(* Logix 5000 project; controller FV vendor 1 type 14 code 217 rev 31.11; software revision 31.00; part 10 of 63 *)
(* tags used below, declared in another part *)
   CWD : CHECKWORD_FLAGS;
   FR_AUDI1 : PlantItem;   // AUDI1
   FR_AUDI1_RawOutput : ALIAS FOR RIO_Rack_2:11:O.Data.30;   // FR_AUDI1
   FR_BEACON1 : PlantItem;   // BEACON1
   FR_BEACON1_RawOutput : ALIAS FOR RIO_Rack_2:11:O.Data.31;   // FR_BEACON1
   FR_data_file_value_to_move : DINT;
   FR_DEFOAM : PlantItem;   // DEFOAM
   FR_DEFOAM_RawOutput : ALIAS FOR RIO_Rack_2:5:O.Data.6;   // FR_DEFOAM
   FR_Delphi_O : DINT[60];
   FR_FV26_VA01 : PlantItem;   // FV26_VA01
   FR_FV26_VA01_RawOutput : ALIAS FOR RIO_Rack_2:11:O.Data.24;   // FR_FV26_VA01
   FR_FV27_VA01 : PlantItem;   // FV27_VA01
   FR_FV27_VA01_RawOutput : ALIAS FOR RIO_Rack_2:11:O.Data.25;   // FR_FV27_VA01
   FR_FV28_V : PlantItem;   // FV28_V
   FR_FV28_V_RawOutput : ALIAS FOR RIO_Rack_2:11:O.Data.20;   // FR_FV28_V
   FR_FV28_VA01 : PlantItem;   // FV28_VA01
   FR_FV28_VA01_RawOutput : ALIAS FOR RIO_Rack_2:11:O.Data.26;   // FR_FV28_VA01
   FR_FV29_VA01 : PlantItem;   // FV29_VA01
   FR_FV29_VA01_RawOutput : ALIAS FOR RIO_Rack_2:11:O.Data.27;   // FR_FV29_VA01
   FR_FV30_VA01 : PlantItem;   // FV30_VA01
   FR_FV30_VA01_RawOutput : ALIAS FOR RIO_Rack_2:11:O.Data.28;   // FR_FV30_VA01
   FR_FV31_VA01 : PlantItem;   // FV31_VA01
   FR_FV31_VA01_RawOutput : ALIAS FOR RIO_Rack_2:11:O.Data.29;   // FR_FV31_VA01
   FR_FVR1_P01 : PlantItem;   // FVR1_P01
   FR_N130 : INT[265];   // FILTRATE Filtrate Return
   FR_N14 : INT[265];   // MVFV CIP Comms to MVFV CIP Un it PLC
   FR_N140 : INT[265];   // CIP
   FR_N160 : INT[265];   // VESSEL Vessel Working Direc tory
   FR_N99 : INT[265];   // COMMENT Comment Lines
   FR_T131 : TIMER[255];   // FILTRATE
   FR_T4 : TIMER[255];   // TIMER
   FR_YC_1 : PlantItem;   // YC_1
   FR_YC_1_RawOutput : ALIAS FOR RIO_Rack_2:11:O.Data.16;   // FR_YC_1
   FR_YC_2 : PlantItem;   // YC_2
   FR_YC_2_RawOutput : ALIAS FOR RIO_Rack_2:11:O.Data.17;   // FR_YC_2
   FR_YP1_CIP : PlantItem;   // YP1_CIP
   FR_YP1_CIP_RawOutput : ALIAS FOR RIO_Rack_2:11:O.Data.21;   // FR_YP1_CIP
   FR_YP2_CIP : PlantItem;   // YP2_CIP
   FR_YP2_CIP_RawOutput : ALIAS FOR RIO_Rack_2:11:O.Data.22;   // FR_YP2_CIP
   FR_YP3_CIP : PlantItem;   // YP3_CIP
   FR_YP3_CIP_RawOutput : ALIAS FOR RIO_Rack_2:11:O.Data.23;   // FR_YP3_CIP
   FT_Filtrate_131_temp_real : REAL;
(* FR_Common, continued *)

ROUTINE FR_Digital_Outputs   (* ladder *)
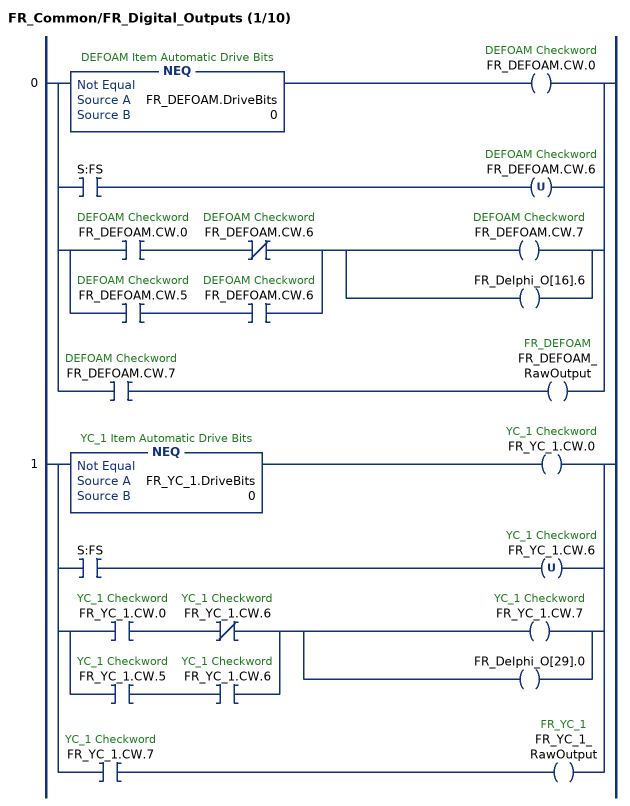
   0: [NEQ(FR_DEFOAM.DriveBits,0) OTE(FR_DEFOAM.CW.0) ,XIC(S:FS) OTU(FR_DEFOAM.CW.6) ,[XIC(FR_DEFOAM.CW.0) XIO(FR_DEFOAM.CW.6) ,XIC(FR_DEFOAM.CW.5) XIC(FR_DEFOAM.CW.6) ] [OTE(FR_DEFOAM.CW.7) ,OTE(FR_Delphi_O[16].6) ] ,XIC(FR_DEFOAM.CW.7) OTE(FR_DEFOAM_RawOutput) ];
   1: [NEQ(FR_YC_1.DriveBits,0) OTE(FR_YC_1.CW.0) ,XIC(S:FS) OTU(FR_YC_1.CW.6) ,[XIC(FR_YC_1.CW.0) XIO(FR_YC_1.CW.6) ,XIC(FR_YC_1.CW.5) XIC(FR_YC_1.CW.6) ] [OTE(FR_YC_1.CW.7) ,OTE(FR_Delphi_O[29].0) ] ,XIC(FR_YC_1.CW.7) OTE(FR_YC_1_RawOutput) ];
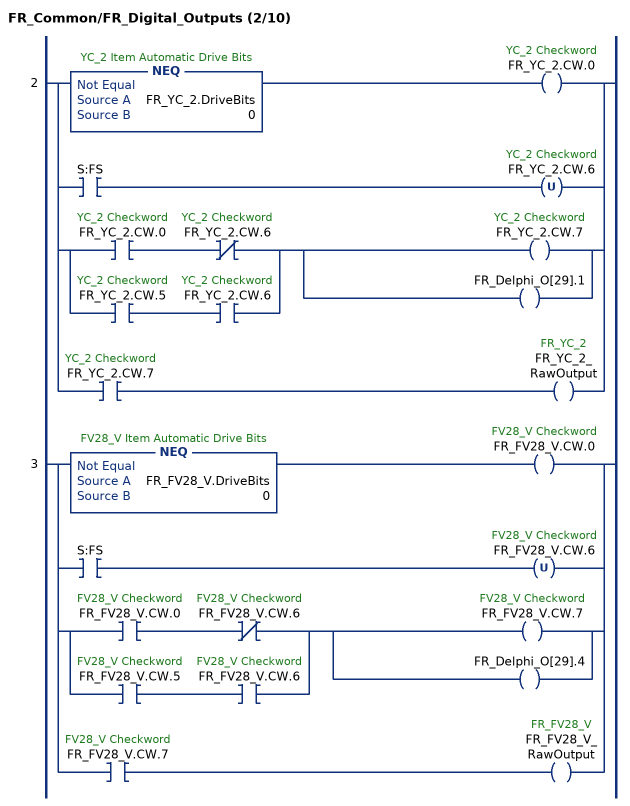
   2: [NEQ(FR_YC_2.DriveBits,0) OTE(FR_YC_2.CW.0) ,XIC(S:FS) OTU(FR_YC_2.CW.6) ,[XIC(FR_YC_2.CW.0) XIO(FR_YC_2.CW.6) ,XIC(FR_YC_2.CW.5) XIC(FR_YC_2.CW.6) ] [OTE(FR_YC_2.CW.7) ,OTE(FR_Delphi_O[29].1) ] ,XIC(FR_YC_2.CW.7) OTE(FR_YC_2_RawOutput) ];
   3: [NEQ(FR_FV28_V.DriveBits,0) OTE(FR_FV28_V.CW.0) ,XIC(S:FS) OTU(FR_FV28_V.CW.6) ,[XIC(FR_FV28_V.CW.0) XIO(FR_FV28_V.CW.6) ,XIC(FR_FV28_V.CW.5) XIC(FR_FV28_V.CW.6) ] [OTE(FR_FV28_V.CW.7) ,OTE(FR_Delphi_O[29].4) ] ,XIC(FR_FV28_V.CW.7) OTE(FR_FV28_V_RawOutput) ];
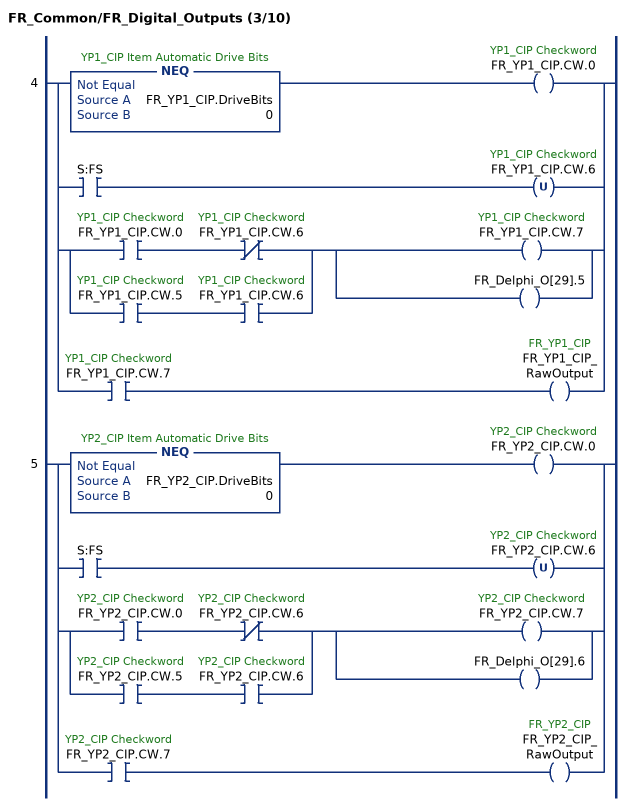
   4: [NEQ(FR_YP1_CIP.DriveBits,0) OTE(FR_YP1_CIP.CW.0) ,XIC(S:FS) OTU(FR_YP1_CIP.CW.6) ,[XIC(FR_YP1_CIP.CW.0) XIO(FR_YP1_CIP.CW.6) ,XIC(FR_YP1_CIP.CW.5) XIC(FR_YP1_CIP.CW.6) ] [OTE(FR_YP1_CIP.CW.7) ,OTE(FR_Delphi_O[29].5) ] ,XIC(FR_YP1_CIP.CW.7) OTE(FR_YP1_CIP_RawOutput) ];
   5: [NEQ(FR_YP2_CIP.DriveBits,0) OTE(FR_YP2_CIP.CW.0) ,XIC(S:FS) OTU(FR_YP2_CIP.CW.6) ,[XIC(FR_YP2_CIP.CW.0) XIO(FR_YP2_CIP.CW.6) ,XIC(FR_YP2_CIP.CW.5) XIC(FR_YP2_CIP.CW.6) ] [OTE(FR_YP2_CIP.CW.7) ,OTE(FR_Delphi_O[29].6) ] ,XIC(FR_YP2_CIP.CW.7) OTE(FR_YP2_CIP_RawOutput) ];
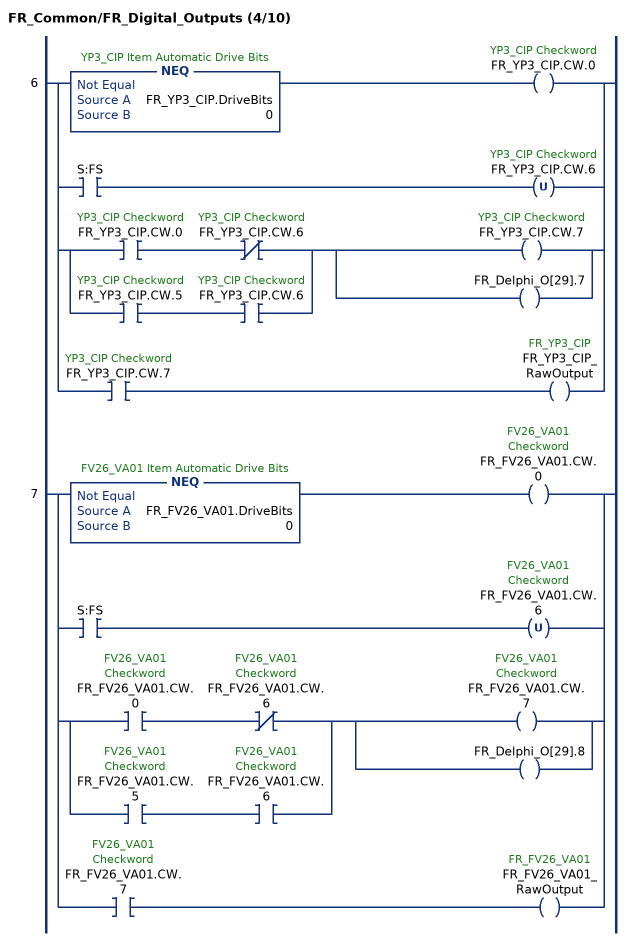
   6: [NEQ(FR_YP3_CIP.DriveBits,0) OTE(FR_YP3_CIP.CW.0) ,XIC(S:FS) OTU(FR_YP3_CIP.CW.6) ,[XIC(FR_YP3_CIP.CW.0) XIO(FR_YP3_CIP.CW.6) ,XIC(FR_YP3_CIP.CW.5) XIC(FR_YP3_CIP.CW.6) ] [OTE(FR_YP3_CIP.CW.7) ,OTE(FR_Delphi_O[29].7) ] ,XIC(FR_YP3_CIP.CW.7) OTE(FR_YP3_CIP_RawOutput) ];
   7: [NEQ(FR_FV26_VA01.DriveBits,0) OTE(FR_FV26_VA01.CW.0) ,XIC(S:FS) OTU(FR_FV26_VA01.CW.6) ,[XIC(FR_FV26_VA01.CW.0) XIO(FR_FV26_VA01.CW.6) ,XIC(FR_FV26_VA01.CW.5) XIC(FR_FV26_VA01.CW.6) ] [OTE(FR_FV26_VA01.CW.7) ,OTE(FR_Delphi_O[29].8) ] ,XIC(FR_FV26_VA01.CW.7) OTE(FR_FV26_VA01_RawOutput) ];
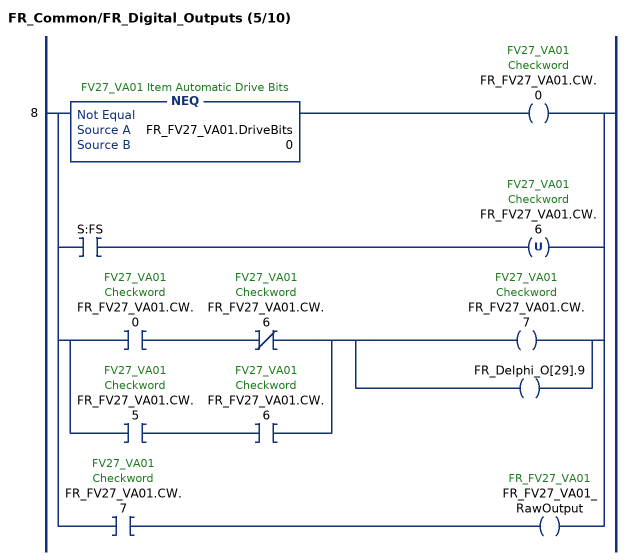
   8: [NEQ(FR_FV27_VA01.DriveBits,0) OTE(FR_FV27_VA01.CW.0) ,XIC(S:FS) OTU(FR_FV27_VA01.CW.6) ,[XIC(FR_FV27_VA01.CW.0) XIO(FR_FV27_VA01.CW.6) ,XIC(FR_FV27_VA01.CW.5) XIC(FR_FV27_VA01.CW.6) ] [OTE(FR_FV27_VA01.CW.7) ,OTE(FR_Delphi_O[29].9) ] ,XIC(FR_FV27_VA01.CW.7) OTE(FR_FV27_VA01_RawOutput) ];
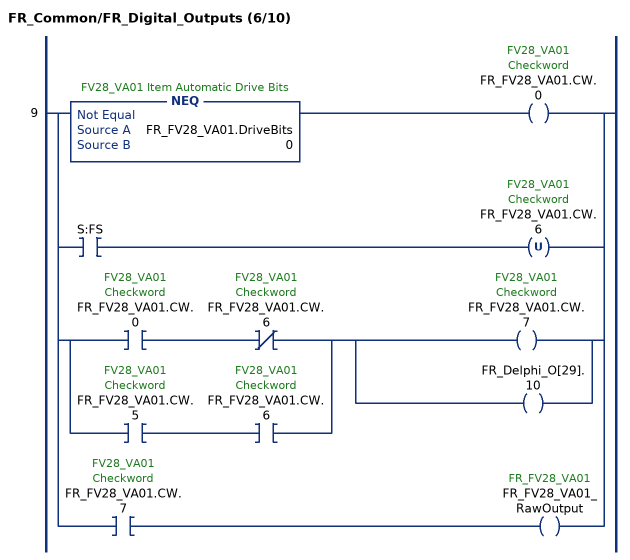
   9: [NEQ(FR_FV28_VA01.DriveBits,0) OTE(FR_FV28_VA01.CW.0) ,XIC(S:FS) OTU(FR_FV28_VA01.CW.6) ,[XIC(FR_FV28_VA01.CW.0) XIO(FR_FV28_VA01.CW.6) ,XIC(FR_FV28_VA01.CW.5) XIC(FR_FV28_VA01.CW.6) ] [OTE(FR_FV28_VA01.CW.7) ,OTE(FR_Delphi_O[29].10) ] ,XIC(FR_FV28_VA01.CW.7) OTE(FR_FV28_VA01_RawOutput) ];
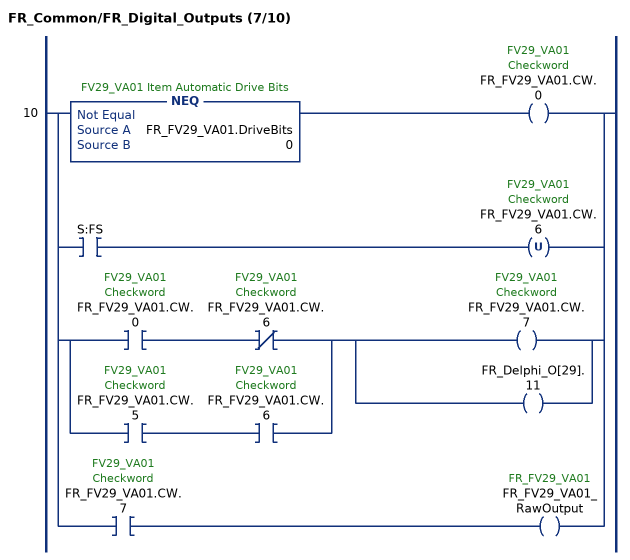
   10: [NEQ(FR_FV29_VA01.DriveBits,0) OTE(FR_FV29_VA01.CW.0) ,XIC(S:FS) OTU(FR_FV29_VA01.CW.6) ,[XIC(FR_FV29_VA01.CW.0) XIO(FR_FV29_VA01.CW.6) ,XIC(FR_FV29_VA01.CW.5) XIC(FR_FV29_VA01.CW.6) ] [OTE(FR_FV29_VA01.CW.7) ,OTE(FR_Delphi_O[29].11) ] ,XIC(FR_FV29_VA01.CW.7) OTE(FR_FV29_VA01_RawOutput) ];
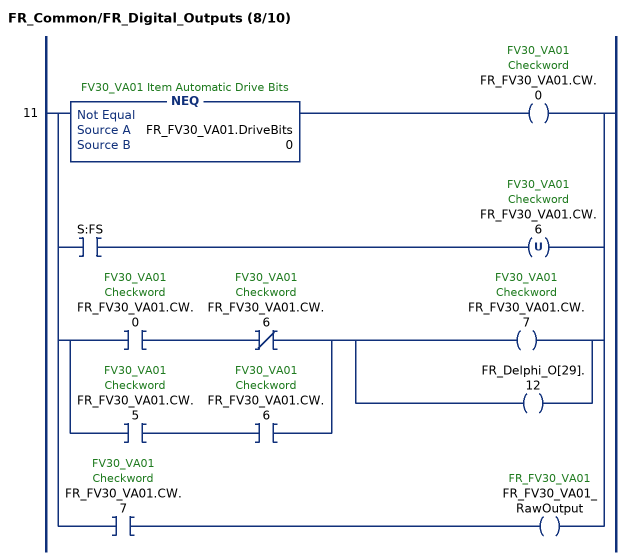
   11: [NEQ(FR_FV30_VA01.DriveBits,0) OTE(FR_FV30_VA01.CW.0) ,XIC(S:FS) OTU(FR_FV30_VA01.CW.6) ,[XIC(FR_FV30_VA01.CW.0) XIO(FR_FV30_VA01.CW.6) ,XIC(FR_FV30_VA01.CW.5) XIC(FR_FV30_VA01.CW.6) ] [OTE(FR_FV30_VA01.CW.7) ,OTE(FR_Delphi_O[29].12) ] ,XIC(FR_FV30_VA01.CW.7) OTE(FR_FV30_VA01_RawOutput) ];
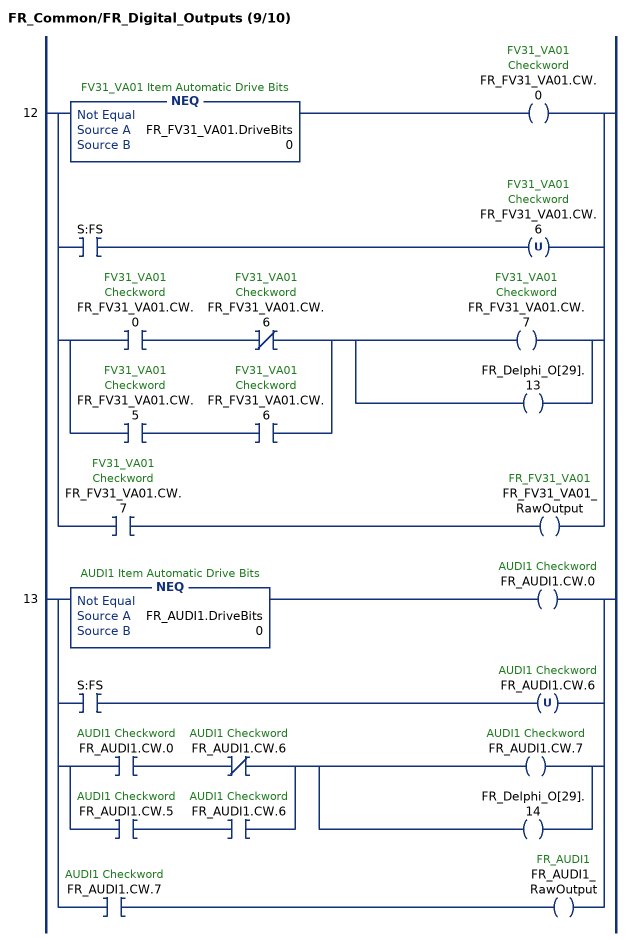
   12: [NEQ(FR_FV31_VA01.DriveBits,0) OTE(FR_FV31_VA01.CW.0) ,XIC(S:FS) OTU(FR_FV31_VA01.CW.6) ,[XIC(FR_FV31_VA01.CW.0) XIO(FR_FV31_VA01.CW.6) ,XIC(FR_FV31_VA01.CW.5) XIC(FR_FV31_VA01.CW.6) ] [OTE(FR_FV31_VA01.CW.7) ,OTE(FR_Delphi_O[29].13) ] ,XIC(FR_FV31_VA01.CW.7) OTE(FR_FV31_VA01_RawOutput) ];
   13: [NEQ(FR_AUDI1.DriveBits,0) OTE(FR_AUDI1.CW.0) ,XIC(S:FS) OTU(FR_AUDI1.CW.6) ,[XIC(FR_AUDI1.CW.0) XIO(FR_AUDI1.CW.6) ,XIC(FR_AUDI1.CW.5) XIC(FR_AUDI1.CW.6) ] [OTE(FR_AUDI1.CW.7) ,OTE(FR_Delphi_O[29].14) ] ,XIC(FR_AUDI1.CW.7) OTE(FR_AUDI1_RawOutput) ];
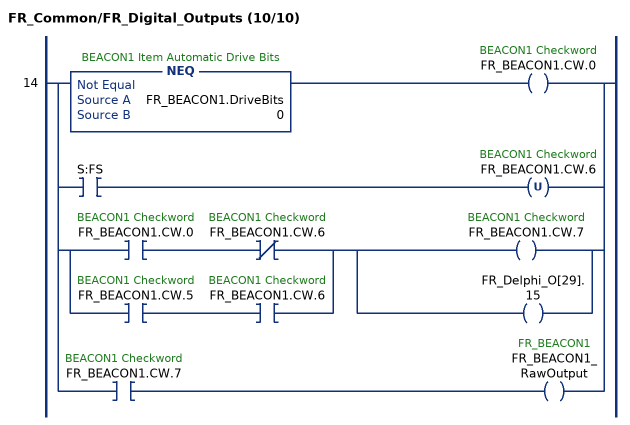
   14: [NEQ(FR_BEACON1.DriveBits,0) OTE(FR_BEACON1.CW.0) ,XIC(S:FS) OTU(FR_BEACON1.CW.6) ,[XIC(FR_BEACON1.CW.0) XIO(FR_BEACON1.CW.6) ,XIC(FR_BEACON1.CW.5) XIC(FR_BEACON1.CW.6) ] [OTE(FR_BEACON1.CW.7) ,OTE(FR_Delphi_O[29].15) ] ,XIC(FR_BEACON1.CW.7) OTE(FR_BEACON1_RawOutput) ];
END_ROUTINE

ROUTINE FR_FILTRATE_131   (* ladder *)
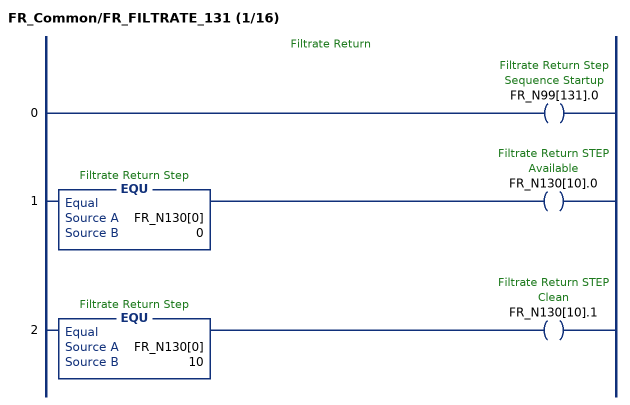
   // Filtrate Return
   0: OTE(FR_N99[131].0);
   1: EQU(FR_N130[0],0)OTE(FR_N130[10].0);
   2: EQU(FR_N130[0],10)OTE(FR_N130[10].1);
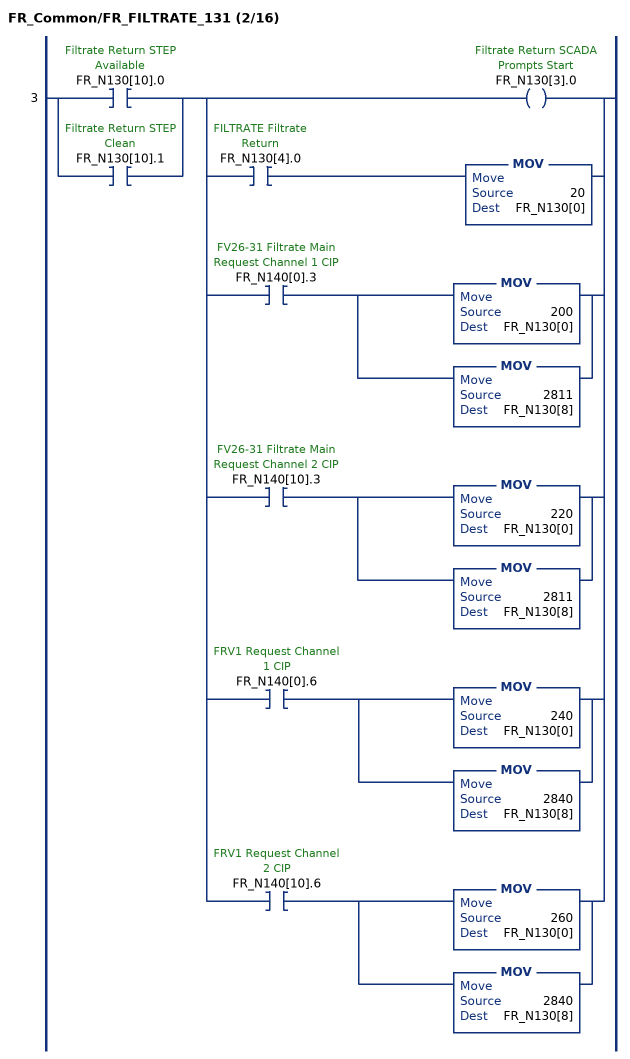
   3: [XIC(FR_N130[10].0) ,XIC(FR_N130[10].1) ][OTE(FR_N130[3].0) ,XIC(FR_N130[4].0) MOV(20,FR_N130[0]) ,XIC(FR_N140[0].3) [MOV(200,FR_N130[0]) ,MOV(2811,FR_N130[8]) ] ,XIC(FR_N140[10].3) [MOV(220,FR_N130[0]) ,MOV(2811,FR_N130[8]) ] ,XIC(FR_N140[0].6) [MOV(240,FR_N130[0]) ,MOV(2840,FR_N130[8]) ] ,XIC(FR_N140[10].6) [MOV(260,FR_N130[0]) ,MOV(2840,FR_N130[8]) ] ];
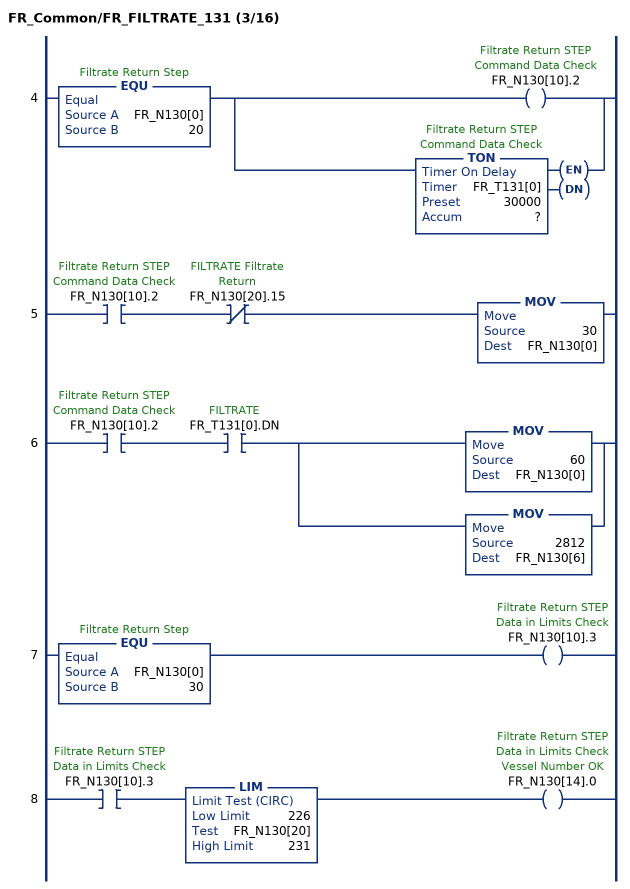
   4: EQU(FR_N130[0],20)[OTE(FR_N130[10].2) ,TON(FR_T131[0],?,?) ];
   5: XIC(FR_N130[10].2)XIO(FR_N130[20].15)MOV(30,FR_N130[0]);
   6: XIC(FR_N130[10].2)XIC(FR_T131[0].DN)[MOV(60,FR_N130[0]) ,MOV(2812,FR_N130[6]) ];
   7: EQU(FR_N130[0],30)OTE(FR_N130[10].3);
   8: XIC(FR_N130[10].3)LIM(226,FR_N130[20],231)OTE(FR_N130[14].0);
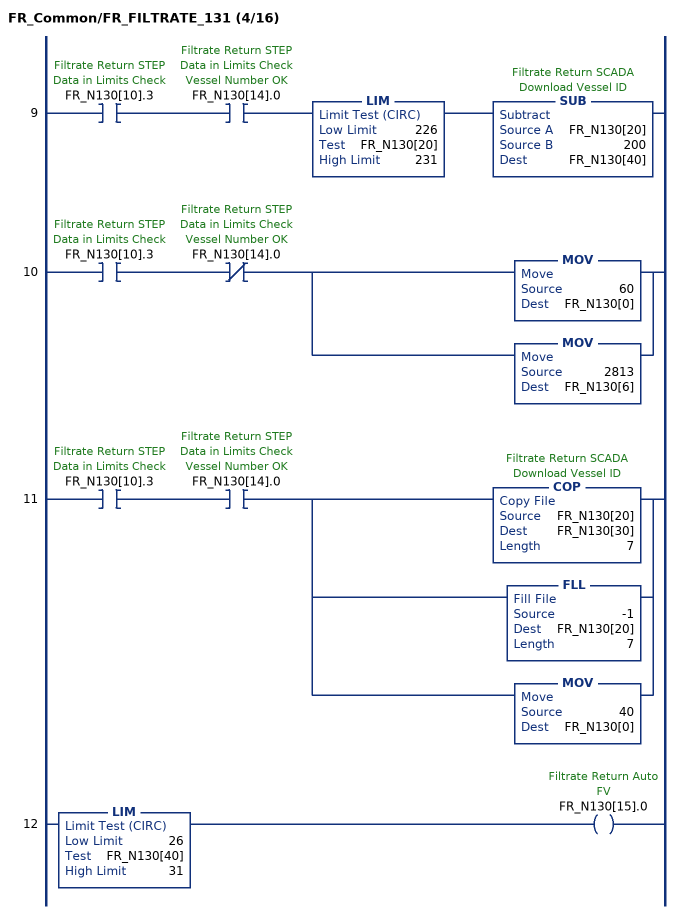
   9: XIC(FR_N130[10].3)XIC(FR_N130[14].0)LIM(226,FR_N130[20],231)SUB(FR_N130[20],200,FR_N130[40]);
   10: XIC(FR_N130[10].3)XIO(FR_N130[14].0)[MOV(60,FR_N130[0]) ,MOV(2813,FR_N130[6]) ];
   11: XIC(FR_N130[10].3)XIC(FR_N130[14].0)[COP(FR_N130[20],FR_N130[30],7) ,FLL(-1,FR_N130[20],7) ,MOV(40,FR_N130[0]) ];
   12: LIM(26,FR_N130[40],31)OTE(FR_N130[15].0);
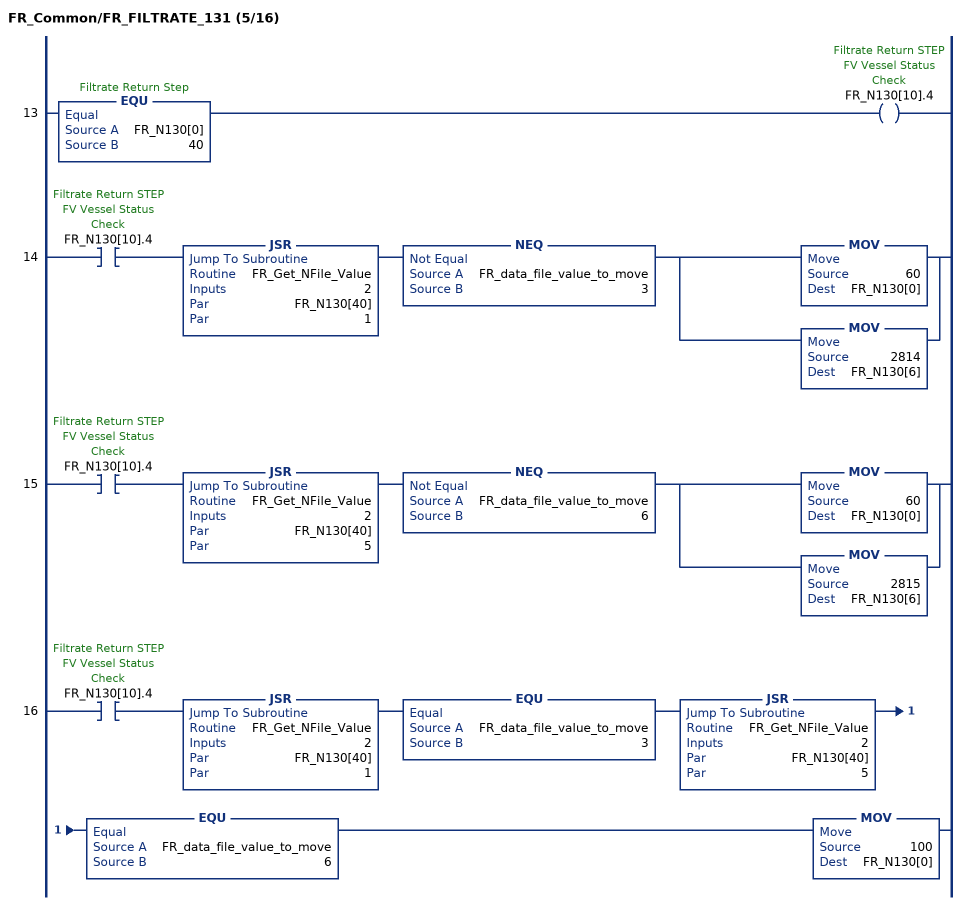
   13: EQU(FR_N130[0],40)OTE(FR_N130[10].4);
   14: XIC(FR_N130[10].4)JSR(FR_Get_NFile_Value,2,FR_N130[40],1)NEQ(FR_data_file_value_to_move,3)[MOV(60,FR_N130[0]) ,MOV(2814,FR_N130[6]) ];
   15: XIC(FR_N130[10].4)JSR(FR_Get_NFile_Value,2,FR_N130[40],5)NEQ(FR_data_file_value_to_move,6)[MOV(60,FR_N130[0]) ,MOV(2815,FR_N130[6]) ];
   16: XIC(FR_N130[10].4)JSR(FR_Get_NFile_Value,2,FR_N130[40],1)EQU(FR_data_file_value_to_move,3)JSR(FR_Get_NFile_Value,2,FR_N130[40],5)EQU(FR_data_file_value_to_move,6)MOV(100,FR_N130[0]);
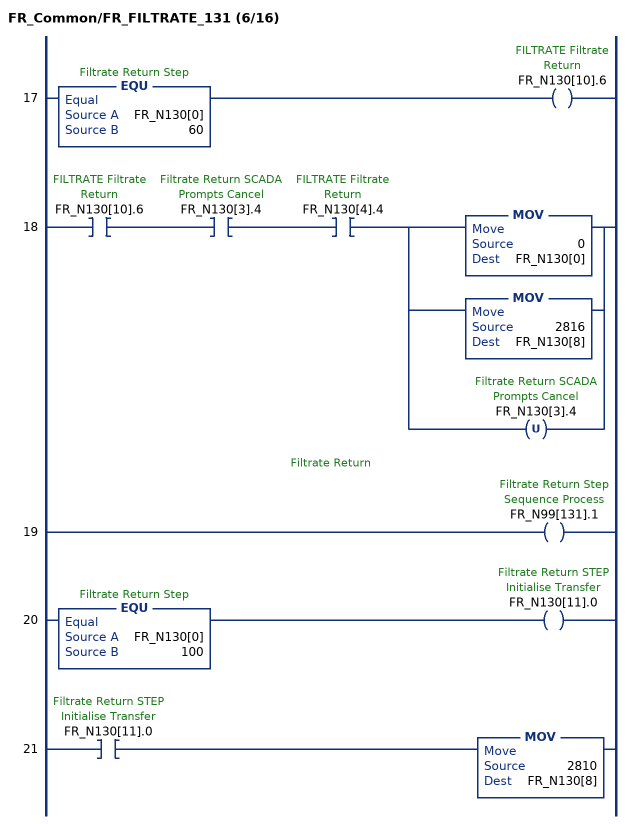
   17: EQU(FR_N130[0],60)OTE(FR_N130[10].6);
   18: XIC(FR_N130[10].6)XIC(FR_N130[3].4)XIC(FR_N130[4].4)[MOV(0,FR_N130[0]) ,MOV(2816,FR_N130[8]) ,OTU(FR_N130[3].4) ];
   // Filtrate Return
   19: OTE(FR_N99[131].1);
   20: EQU(FR_N130[0],100)OTE(FR_N130[11].0);
   21: XIC(FR_N130[11].0)MOV(2810,FR_N130[8]);
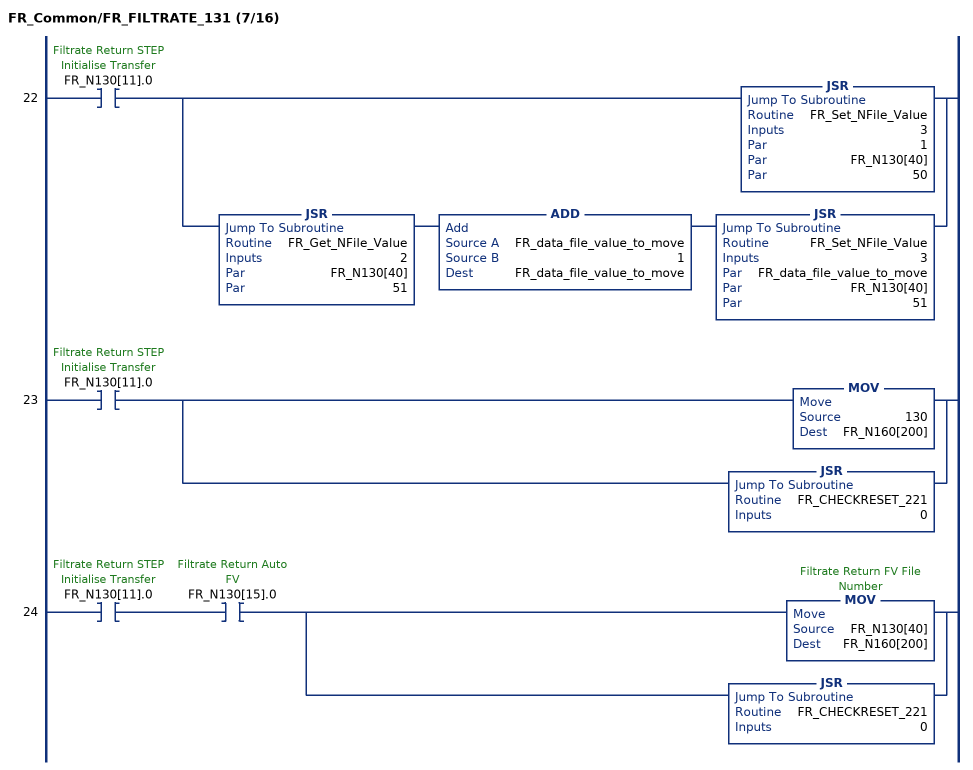
   22: XIC(FR_N130[11].0)[JSR(FR_Set_NFile_Value,3,1,FR_N130[40],50) ,JSR(FR_Get_NFile_Value,2,FR_N130[40],51) ADD(FR_data_file_value_to_move,1,FR_data_file_value_to_move) JSR(FR_Set_NFile_Value,3,FR_data_file_value_to_move,FR_N130[40],51) ];
   23: XIC(FR_N130[11].0)[MOV(130,FR_N160[200]) ,JSR(FR_CHECKRESET_221,0) ];
   24: XIC(FR_N130[11].0)XIC(FR_N130[15].0)[MOV(FR_N130[40],FR_N160[200]) ,JSR(FR_CHECKRESET_221,0) ];
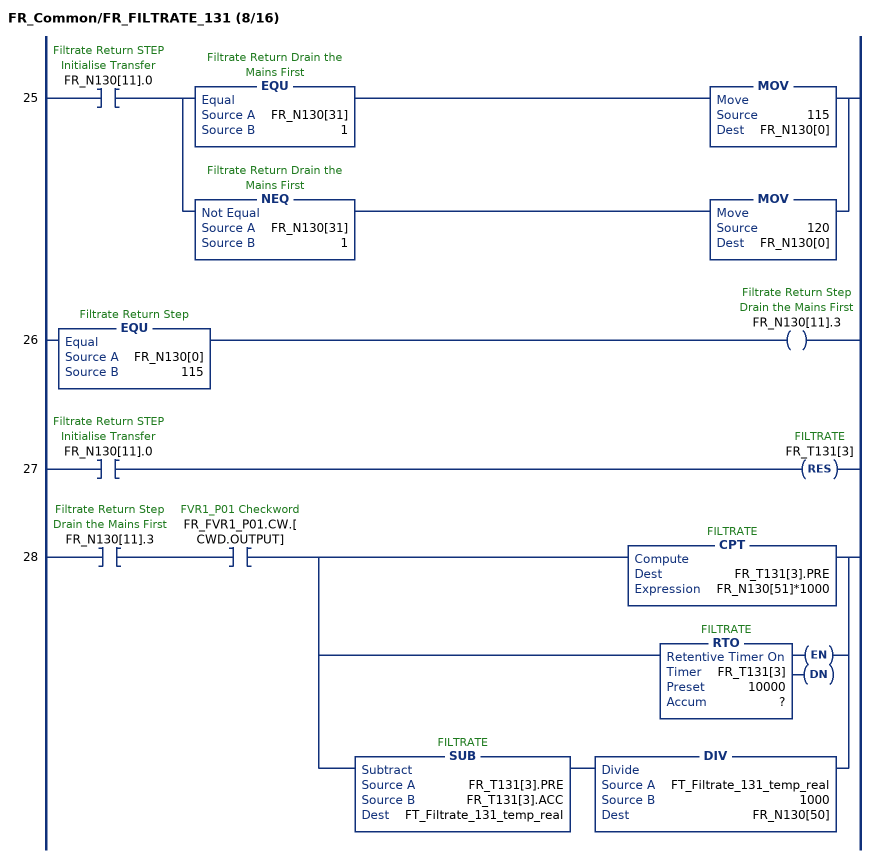
   25: XIC(FR_N130[11].0)[EQU(FR_N130[31],1) MOV(115,FR_N130[0]) ,NEQ(FR_N130[31],1) MOV(120,FR_N130[0]) ];
   26: EQU(FR_N130[0],115)OTE(FR_N130[11].3);
   27: XIC(FR_N130[11].0)RES(FR_T131[3]);
   28: XIC(FR_N130[11].3)XIC(FR_FVR1_P01.CW.[CWD.OUTPUT])[CPT(FR_T131[3].PRE,FR_N130[51]*1000) ,RTO(FR_T131[3],?,?) ,SUB(FR_T131[3].PRE,FR_T131[3].ACC,FT_Filtrate_131_temp_real) DIV(FT_Filtrate_131_temp_real,1000,FR_N130[50]) ];
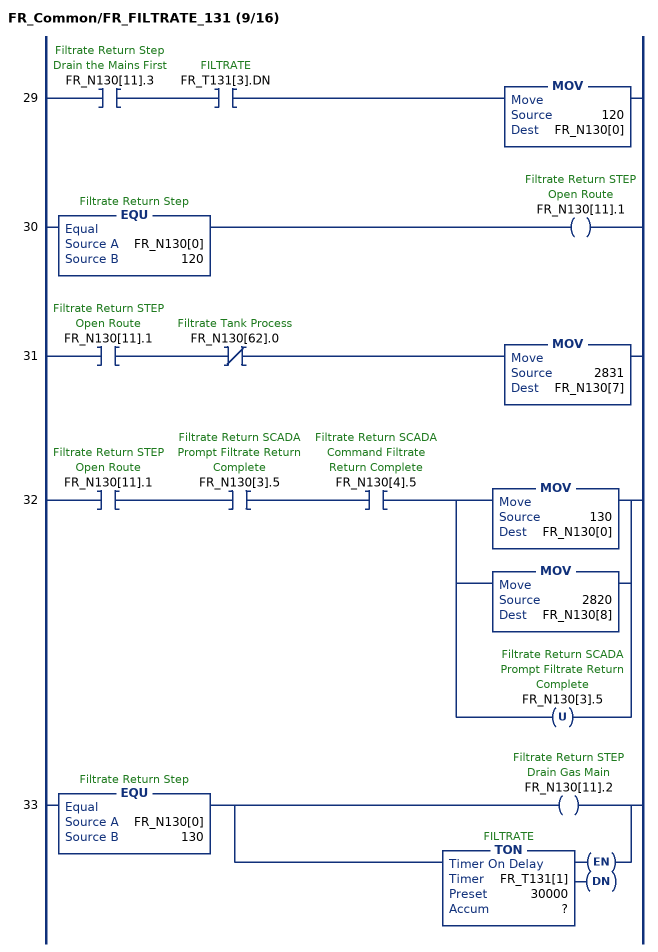
   29: XIC(FR_N130[11].3)XIC(FR_T131[3].DN)MOV(120,FR_N130[0]);
   30: EQU(FR_N130[0],120)OTE(FR_N130[11].1);
   31: XIC(FR_N130[11].1)XIO(FR_N130[62].0)MOV(2831,FR_N130[7]);
   32: XIC(FR_N130[11].1)XIC(FR_N130[3].5)XIC(FR_N130[4].5)[MOV(130,FR_N130[0]) ,MOV(2820,FR_N130[8]) ,OTU(FR_N130[3].5) ];
   33: EQU(FR_N130[0],130)[OTE(FR_N130[11].2) ,TON(FR_T131[1],?,?) ];
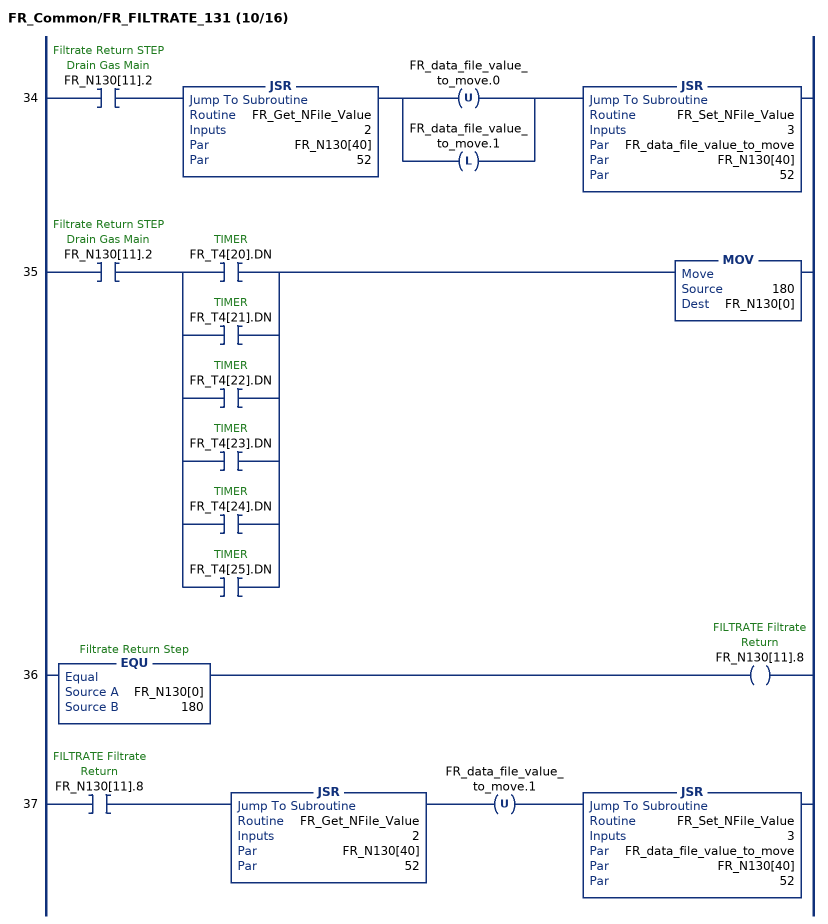
   34: XIC(FR_N130[11].2)JSR(FR_Get_NFile_Value,2,FR_N130[40],52)[OTU(FR_data_file_value_to_move.0) ,OTL(FR_data_file_value_to_move.1) ]JSR(FR_Set_NFile_Value,3,FR_data_file_value_to_move,FR_N130[40],52);
   35: XIC(FR_N130[11].2)[XIC(FR_T4[20].DN) ,XIC(FR_T4[21].DN) ,XIC(FR_T4[22].DN) ,XIC(FR_T4[23].DN) ,XIC(FR_T4[24].DN) ,XIC(FR_T4[25].DN) ]MOV(180,FR_N130[0]);
   36: EQU(FR_N130[0],180)OTE(FR_N130[11].8);
   37: XIC(FR_N130[11].8)JSR(FR_Get_NFile_Value,2,FR_N130[40],52)OTU(FR_data_file_value_to_move.1)JSR(FR_Set_NFile_Value,3,FR_data_file_value_to_move,FR_N130[40],52);
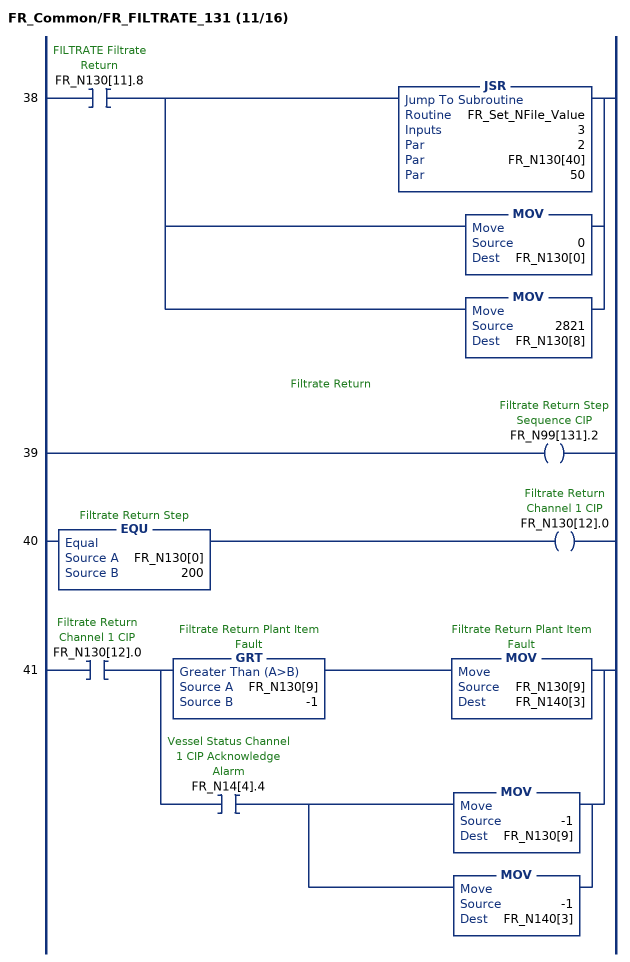
   38: XIC(FR_N130[11].8)[JSR(FR_Set_NFile_Value,3,2,FR_N130[40],50) ,MOV(0,FR_N130[0]) ,MOV(2821,FR_N130[8]) ];
   // Filtrate Return
   39: OTE(FR_N99[131].2);
   40: EQU(FR_N130[0],200)OTE(FR_N130[12].0);
   41: XIC(FR_N130[12].0)[GRT(FR_N130[9],-1) MOV(FR_N130[9],FR_N140[3]) ,XIC(FR_N14[4].4) [MOV(-1,FR_N130[9]) ,MOV(-1,FR_N140[3]) ] ];
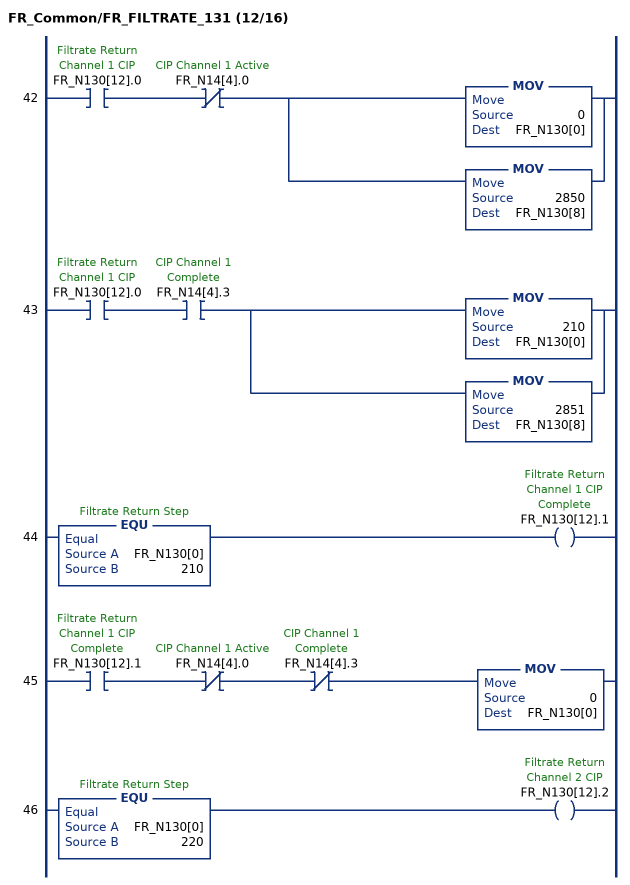
   42: XIC(FR_N130[12].0)XIO(FR_N14[4].0)[MOV(0,FR_N130[0]) ,MOV(2850,FR_N130[8]) ];
   43: XIC(FR_N130[12].0)XIC(FR_N14[4].3)[MOV(210,FR_N130[0]) ,MOV(2851,FR_N130[8]) ];
   44: EQU(FR_N130[0],210)OTE(FR_N130[12].1);
   45: XIC(FR_N130[12].1)XIO(FR_N14[4].0)XIO(FR_N14[4].3)MOV(0,FR_N130[0]);
   46: EQU(FR_N130[0],220)OTE(FR_N130[12].2);
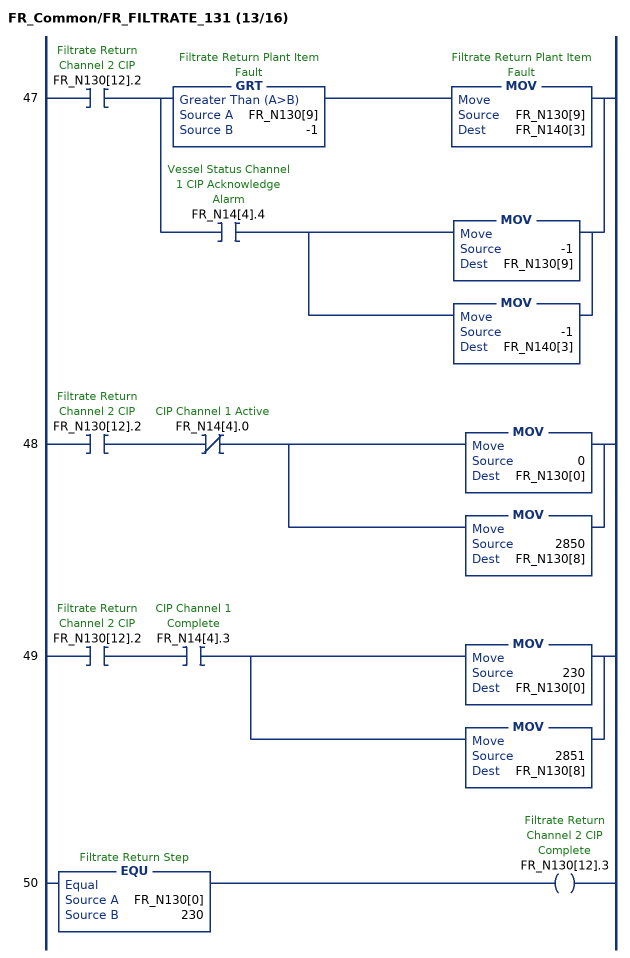
   47: XIC(FR_N130[12].2)[GRT(FR_N130[9],-1) MOV(FR_N130[9],FR_N140[3]) ,XIC(FR_N14[4].4) [MOV(-1,FR_N130[9]) ,MOV(-1,FR_N140[3]) ] ];
   48: XIC(FR_N130[12].2)XIO(FR_N14[4].0)[MOV(0,FR_N130[0]) ,MOV(2850,FR_N130[8]) ];
   49: XIC(FR_N130[12].2)XIC(FR_N14[4].3)[MOV(230,FR_N130[0]) ,MOV(2851,FR_N130[8]) ];
   50: EQU(FR_N130[0],230)OTE(FR_N130[12].3);
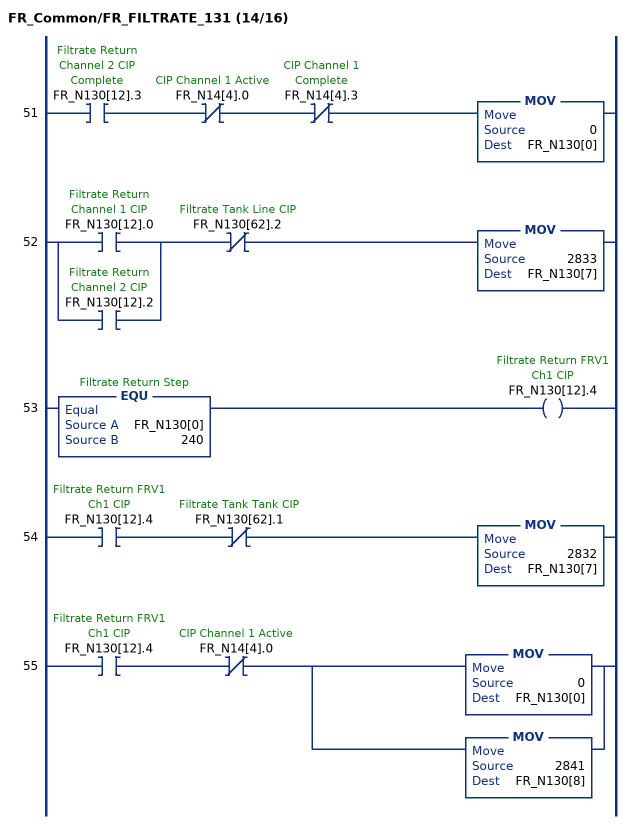
   51: XIC(FR_N130[12].3)XIO(FR_N14[4].0)XIO(FR_N14[4].3)MOV(0,FR_N130[0]);
   52: [XIC(FR_N130[12].0) ,XIC(FR_N130[12].2) ]XIO(FR_N130[62].2)MOV(2833,FR_N130[7]);
   53: EQU(FR_N130[0],240)OTE(FR_N130[12].4);
   54: XIC(FR_N130[12].4)XIO(FR_N130[62].1)MOV(2832,FR_N130[7]);
   55: XIC(FR_N130[12].4)XIO(FR_N14[4].0)[MOV(0,FR_N130[0]) ,MOV(2841,FR_N130[8]) ];
